(* Logix 5000 project; controller _GigaDiscovery vendor 1 type 14 code 244 rev 35.11; software revision 35.03; part 23 of 23 *)
(* tags used below, declared in another part *)
   O_Safety_Valve_Unlock_Left_Block : BOOL;   // Steps 02 to 21
   O_Safety_Valve_Unlock_Right_Block : BOOL;   // Steps 02 to 21
   Proof_Test : Proof_Test;
   No_Sfty : Std_to_Sfty;
   O_RESTRAINTS_Main_Valve : BOOL;   // Main Valve -B40501I
   O_RESTRAINTS_Valve_Lift : BOOL;   // Steps 03 04 05
   Restraints_Cycle : Sequencer;
   RESTRAINTS_Sector : LapBars_Sector[9];
   RESTRAINTS_Sector_Enable_OFF : BOOL;   // ALL RESTRAINTS rack commands OFF
   RESTRAINTS_Sector_Enable_ON : BOOL;   // ALL RESTRAINTS Sector Enable ON
(* S_Restraints_Release, continued *)

ROUTINE _99_Commands   (* ladder *)
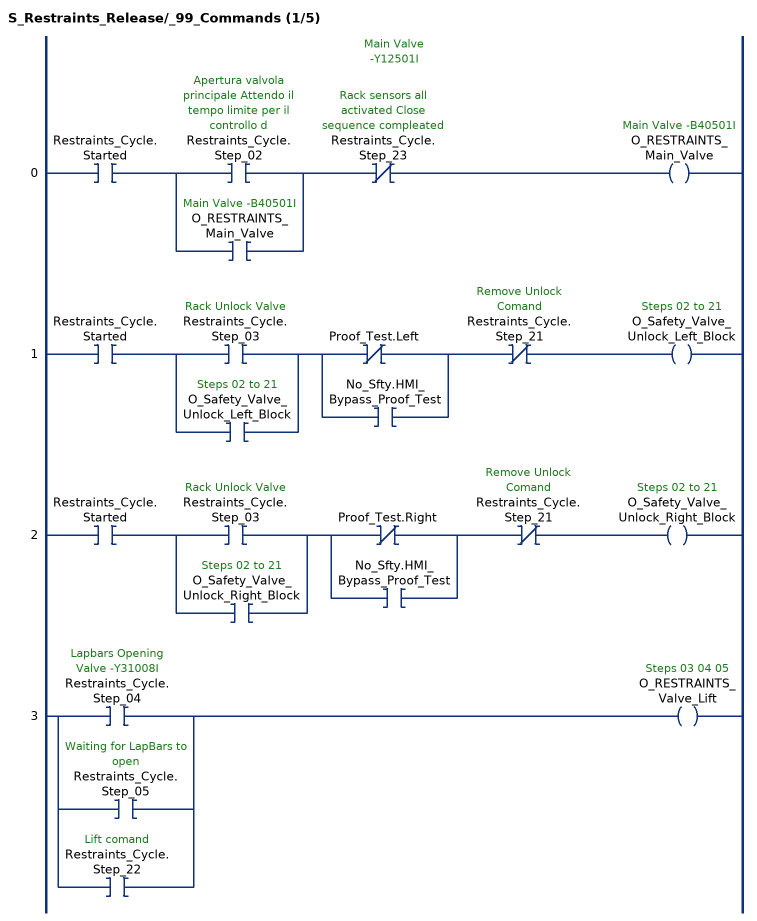
   // Main Valve
   // -Y12501I
   0: XIC(Restraints_Cycle.Started)[XIC(Restraints_Cycle.Step_02) ,XIC(O_RESTRAINTS_Main_Valve) ]XIO(Restraints_Cycle.Step_23)OTE(O_RESTRAINTS_Main_Valve);
   1: XIC(Restraints_Cycle.Started)[XIC(Restraints_Cycle.Step_03) ,XIC(O_Safety_Valve_Unlock_Left_Block) ][XIO(Proof_Test.Left) ,XIC(No_Sfty.HMI_Bypass_Proof_Test) ]XIO(Restraints_Cycle.Step_21)OTE(O_Safety_Valve_Unlock_Left_Block);
   2: XIC(Restraints_Cycle.Started)[XIC(Restraints_Cycle.Step_03) ,XIC(O_Safety_Valve_Unlock_Right_Block) ][XIO(Proof_Test.Right) ,XIC(No_Sfty.HMI_Bypass_Proof_Test) ]XIO(Restraints_Cycle.Step_21)OTE(O_Safety_Valve_Unlock_Right_Block);
   3: [XIC(Restraints_Cycle.Step_04) ,XIC(Restraints_Cycle.Step_05) ,XIC(Restraints_Cycle.Step_22) ]OTE(O_RESTRAINTS_Valve_Lift);
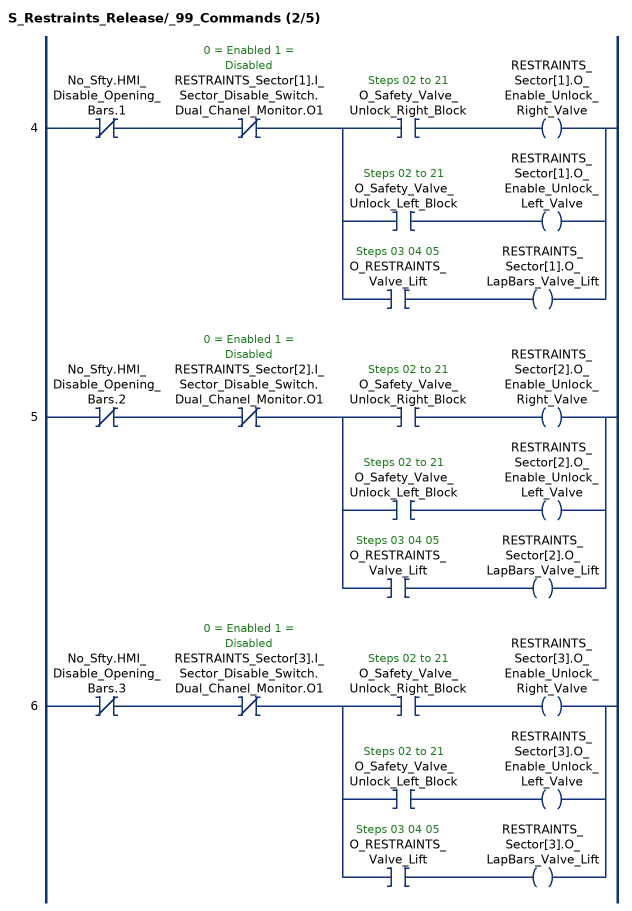
   4: XIO(No_Sfty.HMI_Disable_Opening_Bars.1)XIO(RESTRAINTS_Sector[1].I_Sector_Disable_Switch.Dual_Chanel_Monitor.O1)[XIC(O_Safety_Valve_Unlock_Right_Block) OTE(RESTRAINTS_Sector[1].O_Enable_Unlock_Right_Valve) ,XIC(O_Safety_Valve_Unlock_Left_Block) OTE(RESTRAINTS_Sector[1].O_Enable_Unlock_Left_Valve) ,XIC(O_RESTRAINTS_Valve_Lift) OTE(RESTRAINTS_Sector[1].O_LapBars_Valve_Lift) ];
   5: XIO(No_Sfty.HMI_Disable_Opening_Bars.2)XIO(RESTRAINTS_Sector[2].I_Sector_Disable_Switch.Dual_Chanel_Monitor.O1)[XIC(O_Safety_Valve_Unlock_Right_Block) OTE(RESTRAINTS_Sector[2].O_Enable_Unlock_Right_Valve) ,XIC(O_Safety_Valve_Unlock_Left_Block) OTE(RESTRAINTS_Sector[2].O_Enable_Unlock_Left_Valve) ,XIC(O_RESTRAINTS_Valve_Lift) OTE(RESTRAINTS_Sector[2].O_LapBars_Valve_Lift) ];
   6: XIO(No_Sfty.HMI_Disable_Opening_Bars.3)XIO(RESTRAINTS_Sector[3].I_Sector_Disable_Switch.Dual_Chanel_Monitor.O1)[XIC(O_Safety_Valve_Unlock_Right_Block) OTE(RESTRAINTS_Sector[3].O_Enable_Unlock_Right_Valve) ,XIC(O_Safety_Valve_Unlock_Left_Block) OTE(RESTRAINTS_Sector[3].O_Enable_Unlock_Left_Valve) ,XIC(O_RESTRAINTS_Valve_Lift) OTE(RESTRAINTS_Sector[3].O_LapBars_Valve_Lift) ];
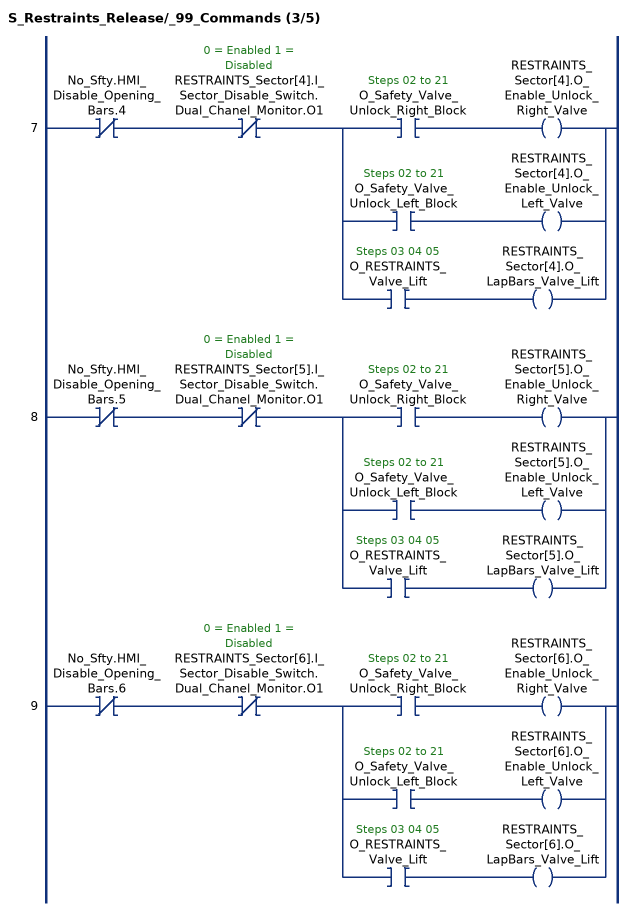
   7: XIO(No_Sfty.HMI_Disable_Opening_Bars.4)XIO(RESTRAINTS_Sector[4].I_Sector_Disable_Switch.Dual_Chanel_Monitor.O1)[XIC(O_Safety_Valve_Unlock_Right_Block) OTE(RESTRAINTS_Sector[4].O_Enable_Unlock_Right_Valve) ,XIC(O_Safety_Valve_Unlock_Left_Block) OTE(RESTRAINTS_Sector[4].O_Enable_Unlock_Left_Valve) ,XIC(O_RESTRAINTS_Valve_Lift) OTE(RESTRAINTS_Sector[4].O_LapBars_Valve_Lift) ];
   8: XIO(No_Sfty.HMI_Disable_Opening_Bars.5)XIO(RESTRAINTS_Sector[5].I_Sector_Disable_Switch.Dual_Chanel_Monitor.O1)[XIC(O_Safety_Valve_Unlock_Right_Block) OTE(RESTRAINTS_Sector[5].O_Enable_Unlock_Right_Valve) ,XIC(O_Safety_Valve_Unlock_Left_Block) OTE(RESTRAINTS_Sector[5].O_Enable_Unlock_Left_Valve) ,XIC(O_RESTRAINTS_Valve_Lift) OTE(RESTRAINTS_Sector[5].O_LapBars_Valve_Lift) ];
   9: XIO(No_Sfty.HMI_Disable_Opening_Bars.6)XIO(RESTRAINTS_Sector[6].I_Sector_Disable_Switch.Dual_Chanel_Monitor.O1)[XIC(O_Safety_Valve_Unlock_Right_Block) OTE(RESTRAINTS_Sector[6].O_Enable_Unlock_Right_Valve) ,XIC(O_Safety_Valve_Unlock_Left_Block) OTE(RESTRAINTS_Sector[6].O_Enable_Unlock_Left_Valve) ,XIC(O_RESTRAINTS_Valve_Lift) OTE(RESTRAINTS_Sector[6].O_LapBars_Valve_Lift) ];
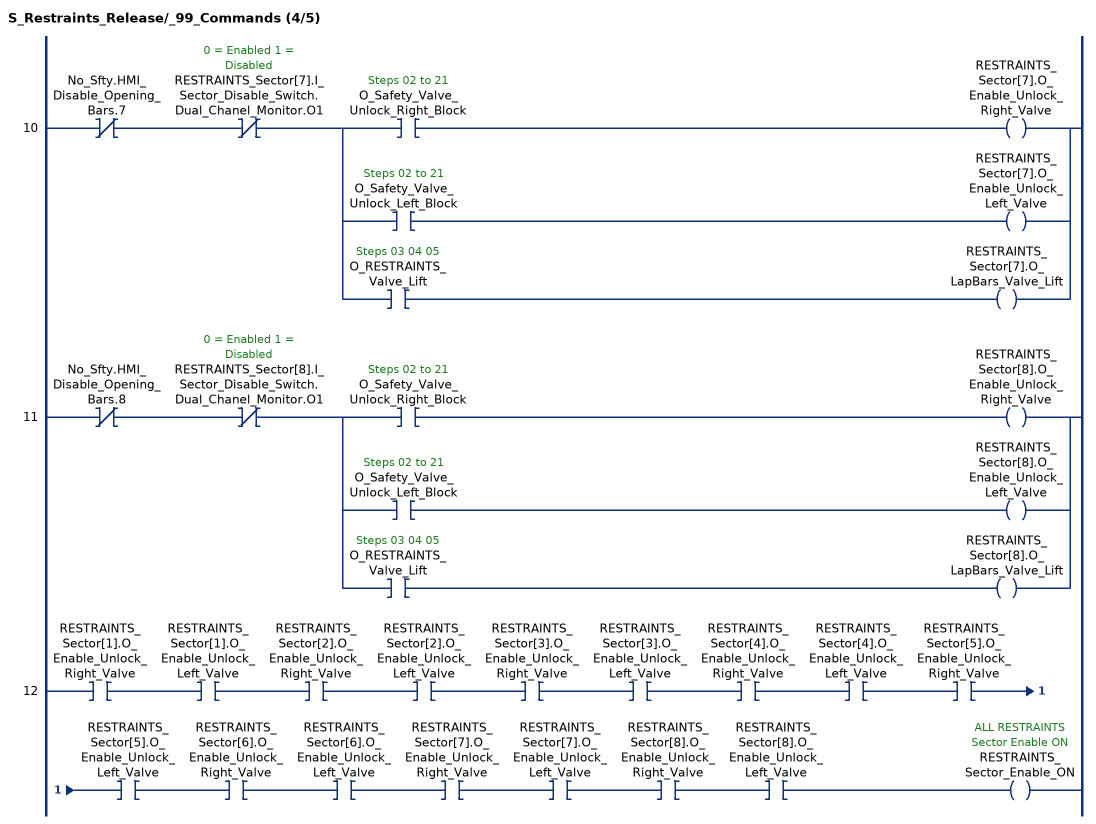
   10: XIO(No_Sfty.HMI_Disable_Opening_Bars.7)XIO(RESTRAINTS_Sector[7].I_Sector_Disable_Switch.Dual_Chanel_Monitor.O1)[XIC(O_Safety_Valve_Unlock_Right_Block) OTE(RESTRAINTS_Sector[7].O_Enable_Unlock_Right_Valve) ,XIC(O_Safety_Valve_Unlock_Left_Block) OTE(RESTRAINTS_Sector[7].O_Enable_Unlock_Left_Valve) ,XIC(O_RESTRAINTS_Valve_Lift) OTE(RESTRAINTS_Sector[7].O_LapBars_Valve_Lift) ];
   11: XIO(No_Sfty.HMI_Disable_Opening_Bars.8)XIO(RESTRAINTS_Sector[8].I_Sector_Disable_Switch.Dual_Chanel_Monitor.O1)[XIC(O_Safety_Valve_Unlock_Right_Block) OTE(RESTRAINTS_Sector[8].O_Enable_Unlock_Right_Valve) ,XIC(O_Safety_Valve_Unlock_Left_Block) OTE(RESTRAINTS_Sector[8].O_Enable_Unlock_Left_Valve) ,XIC(O_RESTRAINTS_Valve_Lift) OTE(RESTRAINTS_Sector[8].O_LapBars_Valve_Lift) ];
   12: XIC(RESTRAINTS_Sector[1].O_Enable_Unlock_Right_Valve)XIC(RESTRAINTS_Sector[1].O_Enable_Unlock_Left_Valve)XIC(RESTRAINTS_Sector[2].O_Enable_Unlock_Right_Valve)XIC(RESTRAINTS_Sector[2].O_Enable_Unlock_Left_Valve)XIC(RESTRAINTS_Sector[3].O_Enable_Unlock_Right_Valve)XIC(RESTRAINTS_Sector[3].O_Enable_Unlock_Left_Valve)XIC(RESTRAINTS_Sector[4].O_Enable_Unlock_Right_Valve)XIC(RESTRAINTS_Sector[4].O_Enable_Unlock_Left_Valve)XIC(RESTRAINTS_Sector[5].O_Enable_Unlock_Right_Valve)XIC(RESTRAINTS_Sector[5].O_Enable_Unlock_Left_Valve)XIC(RESTRAINTS_Sector[6].O_Enable_Unlock_Right_Valve)XIC(RESTRAINTS_Sector[6].O_Enable_Unlock_Left_Valve)XIC(RESTRAINTS_Sector[7].O_Enable_Unlock_Right_Valve)XIC(RESTRAINTS_Sector[7].O_Enable_Unlock_Left_Valve)XIC(RESTRAINTS_Sector[8].O_Enable_Unlock_Right_Valve)XIC(RESTRAINTS_Sector[8].O_Enable_Unlock_Left_Valve)OTE(RESTRAINTS_Sector_Enable_ON);
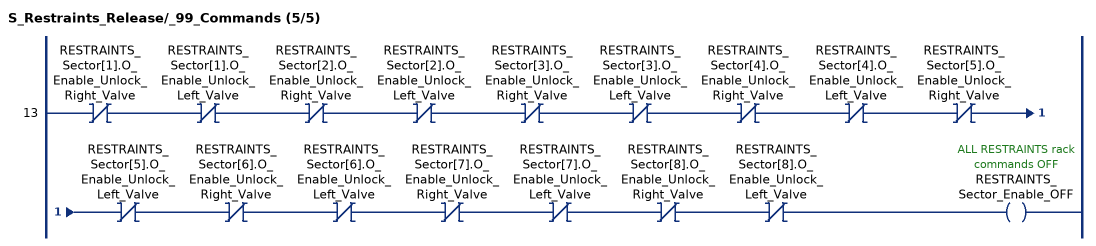
   13: XIO(RESTRAINTS_Sector[1].O_Enable_Unlock_Right_Valve)XIO(RESTRAINTS_Sector[1].O_Enable_Unlock_Left_Valve)XIO(RESTRAINTS_Sector[2].O_Enable_Unlock_Right_Valve)XIO(RESTRAINTS_Sector[2].O_Enable_Unlock_Left_Valve)XIO(RESTRAINTS_Sector[3].O_Enable_Unlock_Right_Valve)XIO(RESTRAINTS_Sector[3].O_Enable_Unlock_Left_Valve)XIO(RESTRAINTS_Sector[4].O_Enable_Unlock_Right_Valve)XIO(RESTRAINTS_Sector[4].O_Enable_Unlock_Left_Valve)XIO(RESTRAINTS_Sector[5].O_Enable_Unlock_Right_Valve)XIO(RESTRAINTS_Sector[5].O_Enable_Unlock_Left_Valve)XIO(RESTRAINTS_Sector[6].O_Enable_Unlock_Right_Valve)XIO(RESTRAINTS_Sector[6].O_Enable_Unlock_Left_Valve)XIO(RESTRAINTS_Sector[7].O_Enable_Unlock_Right_Valve)XIO(RESTRAINTS_Sector[7].O_Enable_Unlock_Left_Valve)XIO(RESTRAINTS_Sector[8].O_Enable_Unlock_Right_Valve)XIO(RESTRAINTS_Sector[8].O_Enable_Unlock_Left_Valve)OTE(RESTRAINTS_Sector_Enable_OFF);
END_ROUTINE

ROUTINE Main   (* ladder *)
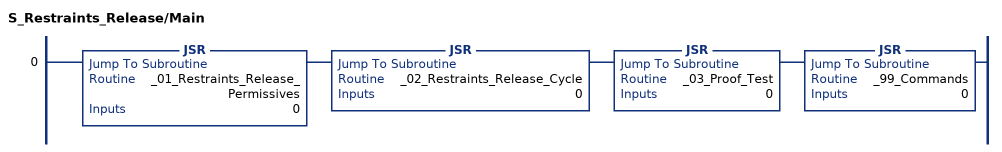
   0: JSR(_01_Restraints_Release_Permissives,0)JSR(_02_Restraints_Release_Cycle,0)JSR(_03_Proof_Test,0)JSR(_99_Commands,0);
END_ROUTINE
END_PROGRAM
